// TIA Portal project "Pesteproject" (V15.1)

(* hardware
DEVICE "S7-1200 station_1"  S7-1200 Station
   slot 0: "Rack_0"  S7-1200 Rack  Rack  V1.0
   slot 1: "PLC_Lines_A_B"  CPU 1212C AC/DC/Rly  6ES7 212-1BE40-0XB0  V4.2
   slot 2: "DI 16x24VDC/DQ 16xRelay_1"  SM 1223 DI16/DQ16 x relay  6ES7 223-1PL32-0XB0  V2.0
   slot 3: "CB 1241 (RS485)"  CB 1241 (RS485)  6ES7 241-1CH30-1XB0  V1.0
   slot 3: "DQ 16xRelay_1"  SM 1222 DQ16 x relay  6ES7 222-1HH32-0XB0  V2.0
DEVICE "S7-1200 station_2"  S7-1200 Station
   slot 0: "Rack_0"  S7-1200 Rack  Rack  V1.0
   slot 1: "PLC_Lines_C"  CPU 1212C AC/DC/Rly  6ES7 212-1BE40-0XB0  V4.2
   slot 2: "DQ 16xRelay_1"  SM 1222 DQ16 x relay  6ES7 222-1HH32-0XB0  V2.0
   slot 3: "CB 1241 (RS485)"  CB 1241 (RS485)  6ES7 241-1CH30-1XB0  V1.0
DEVICE "S71500/ET200MP station_1"  S7-1500 station
   slot 0: "Rail_0"  Rack  6ES7 590-1***0-0AA0
   slot 1: "PLC_1"  CPU 1516-3 PN/DP  6ES7 516-3AN01-0AB0  V2.5
      slot 3: "CPU display_1"  6ES7591-1BA00-0AA0
   slot 2: "DI 16x24VDC BA_1"  DI 16x24VDC BA  6ES7 521-1BH10-0AA0  V1.1
   slot 3: "DI 16x24VDC BA_2"  DI 16x24VDC BA  6ES7 521-1BH10-0AA0  V1.1
*)

// ===== PLC "PLC_Lines_A_B"  CPU 1212C AC/DC/Rly =====

VAR_GLOBAL   // PLC tag table "Default tag table"
   "Phase_Control" AT %I8.0 : Bool;
   "Start_A" AT %I8.7 : Bool;
   "Spare_6" AT %I9.6 : Bool;
   "Spare_7" AT %I9.7 : Bool;
   "Emergency_A" AT %I8.4 : Bool;
   "Fault_A1" AT %I8.1 : Bool;
   "Low_Silo_A1" AT %I0.2 : Bool;
   "Low_Silo_A2" AT %I0.1 : Bool;
   "Low_Silo_B1" AT %I0.7 : Bool;
   "Low_Silo_B2" AT %I0.4 : Bool;
   "High_Silo_A1" AT %I0.3 : Bool;
   "High_Silo_A2" AT %I0.0 : Bool;
   "High_Silo_B1" AT %I0.6 : Bool;
   "High_Silo_B2" AT %I0.5 : Bool;
   "Fault_A2" AT %I9.1 : Bool;
   "Fault_B1" AT %I8.2 : Bool;
   "Fault_B2" AT %I9.2 : Bool;
   "Fault_A3" AT %I9.5 : Bool;
   "Fault_B3" AT %I9.4 : Bool;
   "Emergency_B" AT %I9.3 : Bool;
   "Rel Spare_4" AT %Q2.4 : Bool;
   "Rel Spare_5" AT %Q2.5 : Bool;
   "Rel Spare_6" AT %Q2.6 : Bool;
   "Rel Spare_7" AT %Q2.7 : Bool;
   "Rel Spare_8" AT %Q3.0 : Bool;
   "Rel Spare_9" AT %Q3.1 : Bool;
   "Rel Spare_10" AT %Q3.2 : Bool;
   "Rel Spare_11" AT %Q3.3 : Bool;
   "Rel Spare_12" AT %Q3.4 : Bool;
   "Rel Spare_13" AT %Q3.5 : Bool;
   "Rel Spare_14" AT %Q3.6 : Bool;
   "Rel Spare_15" AT %Q3.7 : Bool;
   "Light_A1" AT %Q2.3 : Bool;
   "Light_A2" AT %Q2.2 : Bool;
   "Light_B1" AT %Q2.1 : Bool;
   "Light_B2" AT %Q2.0 : Bool;
   "Conveyer_A1" AT %Q0.4 : Bool;
   "Conveyer_A2" AT %Q0.5 : Bool;
   "Conveyer_B1" AT %Q9.0 : Bool;
   "Conveyer_B2" AT %Q8.0 : Bool;
   "Pneumatic_A1" AT %Q9.1 : Bool;
   "Pneumatic_A2" AT %Q8.1 : Bool;
   "Pneumatic_B1" AT %Q8.2 : Bool;
   "Pneumatic_B2" AT %Q9.2 : Bool;
   "Conveyer_A3" AT %Q9.5 : Bool;
   "Conveyer_B3_Left" AT %Q9.6 : Bool;
   "Conveyer_B3_Right" AT %Q8.5 : Bool;
   "Tag_1" AT %M10.0 : Bool;
   "Tag_2" AT %M10.1 : Bool;
   "start" AT %M10.2 : Bool;
   "Tag_3" AT %M110.0 : Bool;
   "Tag_10" AT %M110.1 : Bool;
   "Tag_11" AT %M110.2 : Bool;
   "System_Byte" AT %MB1 : Byte;
   "FirstScan" AT %M1.0 : Bool;
   "DiagStatusUpdate" AT %M1.1 : Bool;
   "AlwaysTRUE" AT %M1.2 : Bool;
   "AlwaysFALSE" AT %M1.3 : Bool;
   "Clock_Byte" AT %MB0 : Byte;
   "Clock_10Hz" AT %M0.0 : Bool;
   "Clock_5Hz" AT %M0.1 : Bool;
   "Clock_2.5Hz" AT %M0.2 : Bool;
   "Clock_2Hz" AT %M0.3 : Bool;
   "Clock_1.25Hz" AT %M0.4 : Bool;
   "Clock_1Hz" AT %M0.5 : Bool;
   "Clock_0.625Hz" AT %M0.6 : Bool;
   "Clock_0.5Hz" AT %M0.7 : Bool;
   "Tag_12" AT %M120.1 : Bool;
   "Tag_13" AT %M120.0 : Bool;
   "Tag_14" AT %M120.2 : Bool;
   "Tag_15" AT %MW112 : Word;
   "Tag_16" AT %MW114 : Word;
   "Tag_17" AT %MW122 : Word;
   "Tag_18" AT %MW124 : Word;
   "Tag_4" AT %M1000.0 : Bool;
   "Tag_5" AT %M1000.1 : Bool;
   "Tag_6" AT %MW1002 : Word;
   "Tag_7" AT %M1000.4 : Bool;
   "Tag_8" AT %MW1004 : Word;
   "Tag_9" AT %M1010.0 : Bool;
   "Tag_19" AT %M1010.1 : Bool;
   "Tag_20" AT %M1010.2 : Bool;
   "Tag_21" AT %MW1012 : Word;
   "Tag_22" AT %M1010.4 : Bool;
   "Tag_23" AT %MW1014 : Word;
   "Tag_24" AT %M990.0 : Bool;
   "Tag_25" AT %M990.5 : Bool;
   "Line_A1_Start_Consent" AT %M150.0 : Bool;
   "Line_A1_Run_Consent" AT %M150.1 : Bool;
   "Line_A1_Conveyer_Timer" AT %M150.2 : Bool;
   "A1_Start_Conveyer" AT %M150.3 : Bool;
   "TriggerStartToggleMemory" AT %M150.4 : Bool;
   "Start_A1_Toggle" AT %M150.5 : Bool;
   "TriggerA1ToggleStop" AT %M150.6 : Bool;
   "Conveyer_A1_On" AT %M150.7 : Bool;
   "Conveyer_A1_Off" AT %M151.0 : Bool;
   "Line_A2_Start_Consent" AT %M160.0 : Bool;
   "Line_A2_Run_Consent" AT %M160.1 : Bool;
   "Line_A2_Conveyer_Timer" AT %M160.2 : Bool;
   "A2_Start_Conveyer" AT %M160.3 : Bool;
   "TriggerStopToggleMemoryA2" AT %M160.6 : Bool;
   "TriggerStartToggleMemoryA2" AT %M160.4 : Bool;
   "Start_A2_Toggle" AT %M160.5 : Bool;
   "Conveyer_A2_Off" AT %M161.0 : Bool;
   "Conveyer_A2_On" AT %M160.7 : Bool;
   "Line_B1_Start_Consent" AT %M170.0 : Bool;
   "Line_B1_Run_Consent" AT %M170.1 : Bool;
   "Line_B1_Conveyer_Timer" AT %M170.2 : Bool;
   "B1_Start_Conveyer" AT %M170.3 : Bool;
   "Start_B1_Toggle" AT %M170.5 : Bool;
   "TriggerStartToggleMemoryB1" AT %M170.4 : Bool;
   "TriggerB1ToggleStop" AT %M170.6 : Bool;
   "Conveyer_B1_Off" AT %M171.0 : Bool;
   "Conveyer_B1_On" AT %M170.7 : Bool;
   "Line_B2_Start_Consent" AT %M180.0 : Bool;
   "Line_B2_Run_Consent" AT %M180.1 : Bool;
   "B2_Start_Conveyer" AT %M180.3 : Bool;
   "Line_B2_Conveyer_Timer" AT %M180.2 : Bool;
   "Start_B2_Toggle" AT %M180.5 : Bool;
   "TriggerStartToggleMemoryB2" AT %M180.4 : Bool;
   "TriggerStopToggleMemoryB2" AT %M180.6 : Bool;
   "Conveyer_B2_Off" AT %M181.0 : Bool;
   "Conveyer_B2_On" AT %M180.7 : Bool;
   "Vibrator_A1_On" AT %M151.4 : Bool;
   "Vibrator_A2_On" AT %M161.4 : Bool;
   "Vibrator_B1_On" AT %M171.4 : Bool;
   "Vibrator_B2_On" AT %M181.4 : Bool;
   "A1_Sample_Triger" AT %M151.1 : Bool;
   "Conveyer_A1_OneShut" AT %M151.2 : Bool;
   "Tag_27" AT %M151.3 : Bool;
   "A2_Sample_Triger" AT %M161.1 : Bool;
   "Conveyer_A2_OneShut" AT %M161.2 : Bool;
   "B1_Sample_Triger" AT %M171.1 : Bool;
   "Conveyer_B1_OneShut" AT %M171.2 : Bool;
   "B2_Sample_Triger" AT %M181.1 : Bool;
   "Conveyer_B2_OneShut" AT %M181.2 : Bool;
   "B_Emergency_Flag" AT %M171.3 : Bool;
   "SiloAToggleStart" AT %M190.0 : Bool;
   "SiloBToggleStart" AT %M190.1 : Bool;
   "Conveyor_B3_Left" AT %M200.0 : Bool;
   "Conveyor_B3_Right" AT %M200.1 : Bool;
   "Silo_B_Not_Start_Timer" AT %M190.3 : Bool;
   "Silo_A_Not_Start_Timer" AT %M190.2 : Bool;
   "Conveyor_B3_Start" AT %M190.4 : Bool;
   "Conveyor_A1_Empty_line" AT %M151.5 : Bool;
   "Conveyor_A2_Empty_line" AT %M161.5 : Bool;
   "Conveyor_B1_Empty_line" AT %M171.5 : Bool;
   "Conveyor_B2_Empty_line" AT %M181.5 : Bool;
   "Tag_26" AT %MD156 : DInt;
   "Tag_28" AT %MD166 : DInt;
   "Tag_29" AT %MD176 : DInt;
   "Tag_30" AT %MD186 : DInt;
END_VAR

TYPE "tIMEDATATYPE"
VERSION : 0.1
   STRUCT
      HOUR : String;
      MINUTE : String;
      DAY : String;
      MONTH : String;
      YEAR : String;
   END_STRUCT;
END_TYPE

DATA_BLOCK "ScenarioData"   // DB1
{ S7_Optimized_Access := 'TRUE' }
VERSION : 0.1
   VAR
      DefaultScenario : Int := 1;
      Line_A1_Conveyer_on_Time_Scenario_A : DInt := 2;
      Line_A1_Conveyer_off_Time_Scenario_A : DInt := 3;
      Line_A1_Sampling_Time_Scenario_A : DInt := 4;
      Line_A1_Sampling_OpenTime_Scenario_A : DInt := 5;
      Line_A1_Feeder_Intensity_Scenario_A : Int := 6;
      Line_A1_Duration_Big_Silo_Off_Scenario_A : DInt := 7;
      Line_A1_Feeder_Delay_Before_Stop_Time_Scenario_A : DInt := 8;
      Line_A1_Feeder_Delay_After_Start_Time_Scenario_A : DInt := 9;
      Line_A1_Conveyer_on_Time_Scenario_B : DInt := 10;
      Line_A1_Conveyer_off_Time_Scenario_B : DInt := 11;
      Line_A1_Sampling_Time_Scenario_B : DInt := 12;
      Line_A1_Sampling_OpenTime_Scenario_B : DInt := 13;
      Line_A1_Feeder_Intensity_Scenario_B : Int := 14;
      Line_A1_Duration_Big_Silo_Off_Scenario_B : DInt := 15;
      Line_A1_Feeder_Delay_Before_Stop_Time_Scenario_B : DInt := 16;
      Line_A1_Feeder_Delay_After_Start_Time_Scenario_B : DInt := 17;
      Line_A1_Conveyer_on_Time_Scenario_C : DInt := 18;
      Line_A1_Conveyer_off_Time_Scenario_C : DInt := 19;
      Line_A1_Sampling_Time_Scenario_C : DInt := 20;
      Line_A1_Sampling_OpenTime_Scenario_C : DInt := 21;
      Line_A1_Feeder_Intensity_Scenario_C : Int := 22;
      Line_A1_Duration_Big_Silo_Off_Scenario_C : DInt := 23;
      Line_A1_Feeder_Delay_Before_Stop_Time_Scenario_C : DInt := 24;
      Line_A1_Feeder_Delay_After_Start_Time_Scenario_C : DInt := 25;
      Line_A1_Conveyer_on_Time_Scenario_E : DInt := 26;
      Line_A1_Conveyer_off_Time_Scenario_E : DInt := 27;
      Line_A1_Sampling_Time_Scenario_E : DInt := 28;
      Line_A1_Sampling_OpenTime_Scenario_E : DInt := 29;
      Line_A1_Feeder_Intensity_Scenario_E : Int := 30;
      Line_A1_Duration_Big_Silo_Off_Scenario_E : DInt := 31;
      Line_A1_Feeder_Delay_Before_Stop_Time_Scenario_E : DInt := 32;
      Line_A1_Feeder_Delay_After_Start_Time_Scenario_E : DInt := 33;
      Line_A1_Conveyer_on_Time_Scenario_D : DInt := 34;
      Line_A1_Conveyer_off_Time_Scenario_D : DInt := 35;
      Line_A1_Sampling_Time_Scenario_D : DInt := 36;
      Line_A1_Sampling_OpenTime_Scenario_D : DInt := 37;
      Line_A1_Feeder_Intensity_Scenario_D : Int := 38;
      Line_A1_Duration_Big_Silo_Off_Scenario_D : DInt := 39;
      Line_A1_Feeder_Delay_Before_Stop_Time_Scenario_D : DInt := 40;
      Line_A1_Feeder_Delay_After_Start_Time_Scenario_D : DInt := 41;
      Line_A2_Conveyer_on_Time_Scenario_A : DInt := 42;
      Line_A2_Conveyer_off_Time_Scenario_A : DInt := 43;
      Line_A2_Sampling_Time_Scenario_A : DInt := 44;
      Line_A2_Sampling_OpenTime_Scenario_A : DInt := 45;
      Line_A2_Feeder_Intensity_Scenario_A : Int := 46;
      Line_A2_Duration_Big_Silo_Off_Scenario_A : DInt := 47;
      Line_A2_Feeder_Delay_Before_Stop_Time_Scenario_A : DInt := 48;
      Line_A2_Feeder_Delay_After_Start_Time_Scenario_A : DInt := 49;
      Line_A2_Conveyer_on_Time_Scenario_B : DInt := 50;
      Line_A2_Conveyer_off_Time_Scenario_B : DInt := 51;
      Line_A2_Sampling_Time_Scenario_B : DInt := 52;
      Line_A2_Sampling_OpenTime_Scenario_B : DInt := 53;
      Line_A2_Feeder_Intensity_Scenario_B : Int := 54;
      Line_A2_Duration_Big_Silo_Off_Scenario_B : DInt := 55;
      Line_A2_Feeder_Delay_Before_Stop_Time_Scenario_B : DInt := 56;
      Line_A2_Feeder_Delay_After_Start_Time_Scenario_B : DInt := 57;
      Line_A2_Conveyer_on_Time_Scenario_C : DInt := 58;
      Line_A2_Conveyer_off_Time_Scenario_C : DInt := 59;
      Line_A2_Sampling_Time_Scenario_C : DInt := 60;
      Line_A2_Sampling_OpenTime_Scenario_C : DInt := 61;
      Line_A2_Feeder_Intensity_Scenario_C : Int := 62;
      Line_A2_Duration_Big_Silo_Off_Scenario_C : DInt := 63;
      Line_A2_Feeder_Delay_Before_Stop_Time_Scenario_C : DInt := 64;
      Line_A2_Feeder_Delay_After_Start_Time_Scenario_C : DInt := 65;
      Line_A2_Conveyer_on_Time_Scenario_E : DInt := 66;
      Line_A2_Conveyer_off_Time_Scenario_E : DInt := 67;
      Line_A2_Sampling_Time_Scenario_E : DInt := 68;
      Line_A2_Sampling_OpenTime_Scenario_E : DInt := 69;
      Line_A2_Feeder_Intensity_Scenario_E : Int := 70;
      Line_A2_Duration_Big_Silo_Off_Scenario_E : DInt := 71;
      Line_A2_Feeder_Delay_Before_Stop_Time_Scenario_E : DInt := 72;
      Line_A2_Feeder_Delay_After_Start_Time_Scenario_E : DInt := 73;
      Line_A2_Conveyer_on_Time_Scenario_D : DInt := 74;
      Line_A2_Conveyer_off_Time_Scenario_D : DInt := 75;
      Line_A2_Sampling_Time_Scenario_D : DInt := 76;
      Line_A2_Sampling_OpenTime_Scenario_D : DInt := 77;
      Line_A2_Feeder_Intensity_Scenario_D : Int := 78;
      Line_A2_Duration_Big_Silo_Off_Scenario_D : DInt := 79;
      Line_A2_Feeder_Delay_Before_Stop_Time_Scenario_D : DInt := 80;
      Line_A2_Feeder_Delay_After_Start_Time_Scenario_D : DInt := 81;
      Line_B1_Conveyer_on_Time_Scenario_A : DInt := 82;
      Line_B1_Conveyer_off_Time_Scenario_A : DInt := 83;
      Line_B1_Sampling_Time_Scenario_A : DInt := 84;
      Line_B1_Sampling_OpenTime_Scenario_A : DInt := 85;
      Line_B1_Feeder_Intensity_Scenario_A : Int := 86;
      Line_B1_Duration_Big_Silo_Off_Scenario_A : DInt := 87;
      Line_B1_Feeder_Delay_Before_Stop_Time_Scenario_A : DInt := 88;
      Line_B1_Feeder_Delay_After_Start_Time_Scenario_A : DInt := 89;
      Line_B1_Conveyer_on_Time_Scenario_B : DInt := 90;
      Line_B1_Conveyer_off_Time_Scenario_B : DInt := 91;
      Line_B1_Sampling_Time_Scenario_B : DInt := 92;
      Line_B1_Sampling_OpenTime_Scenario_B : DInt := 93;
      Line_B1_Feeder_Intensity_Scenario_B : Int := 94;
      Line_B1_Duration_Big_Silo_Off_Scenario_B : DInt := 95;
      Line_B1_Feeder_Delay_Before_Stop_Time_Scenario_B : DInt := 96;
      Line_B1_Feeder_Delay_After_Start_Time_Scenario_B : DInt := 97;
      Line_B1_Conveyer_on_Time_Scenario_C : DInt := 98;
      Line_B1_Conveyer_off_Time_Scenario_C : DInt := 99;
      Line_B1_Sampling_Time_Scenario_C : DInt := 100;
      Line_B1_Sampling_OpenTime_Scenario_C : DInt := 101;
      Line_B1_Feeder_Intensity_Scenario_C : Int := 102;
      Line_B1_Duration_Big_Silo_Off_Scenario_C : DInt := 103;
      Line_B1_Feeder_Delay_Before_Stop_Time_Scenario_C : DInt := 104;
      Line_B1_Feeder_Delay_After_Start_Time_Scenario_C : DInt := 105;
      Line_B1_Conveyer_on_Time_Scenario_E : DInt := 106;
      Line_B1_Conveyer_off_Time_Scenario_E : DInt := 107;
      Line_B1_Sampling_Time_Scenario_E : DInt := 108;
      Line_B1_Sampling_OpenTime_Scenario_E : DInt := 109;
      Line_B1_Feeder_Intensity_Scenario_E : Int := 110;
      Line_B1_Duration_Big_Silo_Off_Scenario_E : DInt := 111;
      Line_B1_Feeder_Delay_Before_Stop_Time_Scenario_E : DInt := 112;
      Line_B1_Feeder_Delay_After_Start_Time_Scenario_E : DInt := 113;
      Line_B1_Conveyer_on_Time_Scenario_D : DInt := 114;
      Line_B1_Conveyer_off_Time_Scenario_D : DInt := 115;
      Line_B1_Sampling_Time_Scenario_D : DInt := 116;
      Line_B1_Sampling_OpenTime_Scenario_D : DInt := 117;
      Line_B1_Feeder_Intensity_Scenario_D : Int := 118;
      Line_B1_Duration_Big_Silo_Off_Scenario_D : DInt := 119;
      Line_B1_Feeder_Delay_Before_Stop_Time_Scenario_D : DInt := 120;
      Line_B1_Feeder_Delay_After_Start_Time_Scenario_D : DInt := 121;
      Line_B2_Conveyer_on_Time_Scenario_A : DInt := 122;
      Line_B2_Conveyer_off_Time_Scenario_A : DInt := 123;
      Line_B2_Sampling_Time_Scenario_A : DInt := 124;
      Line_B2_Sampling_OpenTime_Scenario_A : DInt := 125;
      Line_B2_Feeder_Intensity_Scenario_A : Int := 126;
      Line_B2_Duration_Big_Silo_Off_Scenario_A : DInt := 127;
      Line_B2_Feeder_Delay_Before_Stop_Time_Scenario_A : DInt := 128;
      Line_B2_Feeder_Delay_After_Start_Time_Scenario_A : DInt := 129;
      Line_B2_Conveyer_on_Time_Scenario_B : DInt := 130;
      Line_B2_Conveyer_off_Time_Scenario_B : DInt := 131;
      Line_B2_Sampling_Time_Scenario_B : DInt := 132;
      Line_B2_Sampling_OpenTime_Scenario_B : DInt := 133;
      Line_B2_Feeder_Intensity_Scenario_B : Int := 134;
      Line_B2_Duration_Big_Silo_Off_Scenario_B : DInt := 135;
      Line_B2_Feeder_Delay_Before_Stop_Time_Scenario_B : DInt := 136;
      Line_B2_Feeder_Delay_After_Start_Time_Scenario_B : DInt := 137;
      Line_B2_Conveyer_on_Time_Scenario_C : DInt := 138;
      Line_B2_Conveyer_off_Time_Scenario_C : DInt := 139;
      Line_B2_Sampling_Time_Scenario_C : DInt := 140;
      Line_B2_Sampling_OpenTime_Scenario_C : DInt := 141;
      Line_B2_Feeder_Intensity_Scenario_C : Int := 142;
      Line_B2_Duration_Big_Silo_Off_Scenario_C : DInt := 143;
      Line_B2_Feeder_Delay_Before_Stop_Time_Scenario_C : DInt := 144;
      Line_B2_Feeder_Delay_After_Start_Time_Scenario_C : DInt := 145;
      Line_B2_Conveyer_on_Time_Scenario_E : DInt := 146;
      Line_B2_Conveyer_off_Time_Scenario_E : DInt := 147;
      Line_B2_Sampling_Time_Scenario_E : DInt := 148;
      Line_B2_Sampling_OpenTime_Scenario_E : DInt := 149;
      Line_B2_Feeder_Intensity_Scenario_E : Int := 150;
      Line_B2_Duration_Big_Silo_Off_Scenario_E : DInt := 151;
      Line_B2_Feeder_Delay_Before_Stop_Time_Scenario_E : DInt := 152;
      Line_B2_Feeder_Delay_After_Start_Time_Scenario_E : DInt := 153;
      Line_B2_Conveyer_on_Time_Scenario_D : DInt := 154;
      Line_B2_Conveyer_off_Time_Scenario_D : DInt := 155;
      Line_B2_Sampling_Time_Scenario_D : DInt := 156;
      Line_B2_Sampling_OpenTime_Scenario_D : DInt := 157;
      Line_B2_Feeder_Intensity_Scenario_D : Int := 158;
      Line_B2_Duration_Big_Silo_Off_Scenario_D : DInt := 159;
      Line_B2_Feeder_Delay_Before_Stop_Time_Scenario_D : DInt := 160;
      Line_B2_Feeder_Delay_After_Start_Time_Scenario_D : DInt := 161;
      Line_A1_Empty_Line_Time_Scenario_A : DInt := 162;
      Line_A2_Empty_Line_Time_Scenario_A : DInt := 163;
      Line_B1_Empty_Line_Time_Scenario_A : DInt := 164;
      Line_B2_Empty_Line_Time_Scenario_A : DInt := 165;
      Line_A1_Empty_Line_Time_Scenario_B : DInt := 166;
      Line_A2_Empty_Line_Time_Scenario_B : DInt := 167;
      Line_B1_Empty_Line_Time_Scenario_B : DInt := 168;
      Line_B2_Empty_Line_Time_Scenario_B : DInt := 169;
      Line_A1_Empty_Line_Time_Scenario_C : DInt := 170;
      Line_A2_Empty_Line_Time_Scenario_C : DInt := 171;
      Line_B1_Empty_Line_Time_Scenario_C : DInt := 172;
      Line_B2_Empty_Line_Time_Scenario_C : DInt := 173;
      Line_A1_Empty_Line_Time_Scenario_D : DInt := 174;
      Line_A2_Empty_Line_Time_Scenario_D : DInt := 175;
      Line_B1_Empty_Line_Time_Scenario_D : DInt := 176;
      Line_B2_Empty_Line_Time_Scenario_D : DInt := 177;
      Line_A1_Empty_Line_Time_Scenario_E : DInt := 178;
      Line_A2_Empty_Line_Time_Scenario_E : DInt := 179;
      Line_B1_Empty_Line_Time_Scenario_E : DInt := 180;
      Line_B2_Empty_Line_Time_Scenario_E : DInt := 181;
   END_VAR
BEGIN
END_DATA_BLOCK

DATA_BLOCK "Conveyer B1_DB"   // DB5
{ S7_Optimized_Access := 'TRUE' }
VERSION : 0.1
// stored: InstanceOfName Conveyer B1
"Conveyer B1"
BEGIN
END_DATA_BLOCK

DATA_BLOCK "ModbusDataSendToFeeders"   // DB7
{ S7_Optimized_Access := 'FALSE' }
VERSION : 0.1
   VAR
      dataforsend : Array[0..3] of Int;
   END_VAR
BEGIN
   dataforsend[0] := 0;
   dataforsend[1] := 0;
   dataforsend[2] := 0;
   dataforsend[3] := 0;
END_DATA_BLOCK

DATA_BLOCK "Conveyer A1_DB"   // DB12
{ S7_Optimized_Access := 'TRUE' }
VERSION : 0.1
// stored: InstanceOfName Conveyer A1
"Conveyer A1"
BEGIN
END_DATA_BLOCK

DATA_BLOCK "Conveyer A2_DB"   // DB13
{ S7_Optimized_Access := 'TRUE' }
VERSION : 0.1
// stored: InstanceOfName Conveyer A2
"Conveyer A2"
BEGIN
END_DATA_BLOCK

DATA_BLOCK "Conveyer B1_DB_1"   // DB17
{ S7_Optimized_Access := 'TRUE' }
VERSION : 0.1
// stored: InstanceOfName Conveyer B1
"Conveyer B1"
BEGIN
END_DATA_BLOCK

DATA_BLOCK "Conveyer B2_DB"   // DB18
{ S7_Optimized_Access := 'TRUE' }
VERSION : 0.1
// stored: InstanceOfName Conveyer B2
"Conveyer B2"
BEGIN
END_DATA_BLOCK

DATA_BLOCK "Vibrator A1_DB"   // DB19
{ S7_Optimized_Access := 'TRUE' }
VERSION : 0.1
// stored: InstanceOfName Vibrator A1
"Vibrator A1"
BEGIN
END_DATA_BLOCK

DATA_BLOCK "Vibrator A2_DB"   // DB20
{ S7_Optimized_Access := 'TRUE' }
VERSION : 0.1
// stored: InstanceOfName Vibrator A2
"Vibrator A2"
BEGIN
END_DATA_BLOCK

DATA_BLOCK "Vibrator B1_DB"   // DB21
{ S7_Optimized_Access := 'TRUE' }
VERSION : 0.1
// stored: InstanceOfName Vibrator B1
"Vibrator B1"
BEGIN
END_DATA_BLOCK

DATA_BLOCK "Vibrator B2_DB"   // DB22
{ S7_Optimized_Access := 'TRUE' }
VERSION : 0.1
// stored: InstanceOfName Vibrator B2
"Vibrator B2"
BEGIN
END_DATA_BLOCK

DATA_BLOCK "Web_Send"   // DB23
{ S7_Optimized_Access := 'TRUE' }
VERSION : 0.1
   VAR
      "time" : DTL;
      ModbusDone : Bool;
      ModbusStatus : Word;
      A1_Scenario_Type : Int := 2;
      A2_Scenario_Type : Int := 1;
      B1_Scenario_Type : Int := 1;
      B2_Scenario_Type : Int := 1;
      A_Emergency : Bool;
      B_Emergency : Bool;
      A1_Fault : Bool;
      A2_Fault : Bool;
      B1_Fault : Bool;
      B2_Fault : Bool;
      A3_Fault : Bool;
      B3_Fault : Bool;
      A1_Silo_Low : Bool;
      A2_Silo_Low : Bool;
      B1_Silo_Low : Bool;
      B2_Silo_Low : Bool;
      A1_Conveyer : Bool;
      A2_Conveyer : Bool;
      B1_Conveyer : Bool;
      B2_Conveyer : Bool;
      A3_Conveyor : Bool;
      B3_Left_Conveyer : Bool;
      A1_Silo_High : Bool;
      A2_Silo_High : Bool;
      B1_Silo_High : Bool;
      B2_Silo_High : Bool;
      A1_Sample : Bool;
      A2_Sample : Bool;
      B1_Sample : Bool;
      B2_Sample : Bool;
      A1_Running_Duration : Time;
      A1_Pause_Duration : Time;
      A1_Feeder_Vibration_Intensity : Int;
      A1_Ruuning_Online : Time;
      A1_Pause_Online : Time;
      A1_Sample_Interval : Time;
      A1_Sample_Duration : Time;
      A1_Sample_Online : Time;
      A1_Enable : Bool;
      A1_Start : Bool;
      A1_Big_Silo : Bool;
      B1_Running_Duration : Time;
      B1_Pause_Duration : Time;
      B1_Feeder_Vibration_Intensity : Int;
      B1_Ruuning_Online : Time;
      B1_Pause_Online : Time;
      B1_Sample_Interval : Time;
      B1_Sample_Duration : Time;
      B1_Sample_Online : Time;
      B1_Enable : Bool;
      B1_Start : Bool;
      B1_Big_Silo : Bool;
      A2_Running_Duration : Time;
      A2_Pause_Duration : Time;
      A2_Feeder_Vibration_Intensity : Int;
      A2_Ruuning_Online : Time;
      A2_Pause_Online : Time;
      A2_Sample_Interval : Time;
      A2_Sample_Duration : Time;
      A2_Sample_Online : Time;
      A2_Enable : Bool;
      A2_Start : Bool;
      A2_Big_Silo : Bool;
      B2_Running_Duration : Time;
      B2_Pause_Duration : Time;
      B2_Feeder_Vibration_Intensity : Int;
      B2_Ruuning_Online : Time;
      B2_Pause_Online : Time;
      B2_Sample_Interval : Time;
      B2_Sample_Duration : Time;
      B2_Sample_Online : Time;
      B2_Enable : Bool;
      B2_Start : Bool;
      B2_Big_Silo : Bool;
      A1_Manual : Bool;
      A2_Manual : Bool;
      B1_Manual : Bool;
      B2_Manual : Bool;
      A1_Feeder : Bool;
      A2_Feeder : Bool;
      B1_Feeder : Bool;
      B2_Feeder : Bool;
      A1_Duration_Big_Silo_Stop_Time : Time;
      A2_Duration_Big_Silo_Stop_Time : Time;
      B1_Duration_Big_Silo_Stop_Time : Time;
      B2_Duration_Big_Silo_Stop_Time : Time;
      A1_Empty_Line_Time : Time;
      A2_Empty_Line_Time : Time;
      B1_Empty_Line_Time : Time;
      B2_Empty_Line_Time : Time;
      A1_Feeder_Delay_After_Start_Time : Time;
      A2_Feeder_Delay_After_Start_Time : Time;
      B1_Feeder_Delay_After_Start_Time : Time;
      B2_Feeder_Delay_After_Start_Time : Time;
      A1_Feeder_Delay_Before_Stop_Time : Time;
      A2_Feeder_Delay_Before_Stop_Time : Time;
      B1_Feeder_Delay_Before_Stop_Time : Time;
      B2_Feeder_Delay_Before_Stop_Time : Time;
      A1_Feeder_Delay_Time : Time;
      A1_Feeder_Delay_Time_1 : Time;
      A1_Feeder_Delay_Time_2 : Time;
      A1_Feeder_Delay_Time_3 : Time;
      B3_Conveyor : Bool;
   END_VAR
BEGIN
END_DATA_BLOCK

DATA_BLOCK "ConveyerA3_B3_DB"   // DB32
{ S7_Optimized_Access := 'TRUE' }
VERSION : 0.1
// stored: InstanceOfName ConveyerA3_B3
"ConveyerA3_B3"
BEGIN
END_DATA_BLOCK

DATA_BLOCK "Sample_A_DB"   // DB33
{ S7_Optimized_Access := 'TRUE' }
VERSION : 0.1
// stored: InstanceOfName Sample
"Sample"
BEGIN
END_DATA_BLOCK

DATA_BLOCK "Silo_Big_A-B_DB"   // DB34
{ S7_Optimized_Access := 'TRUE' }
VERSION : 0.1
// stored: InstanceOfName Silo_Big_A-B
"Silo_Big_A-B"
BEGIN
END_DATA_BLOCK

DATA_BLOCK "Web_Recieve"   // DB45
{ S7_Optimized_Access := 'FALSE' }
VERSION : 0.1
   VAR
      Line_A1_Save_Data : Bool;
      Line_A1_Save_Data_Advance : Bool;
      Line_A1_Start : Bool;
      Line_A1_Enable : Bool := 0;
      Line_A1_Conveyer_on_Time : Time := T#26MS;
      Line_A1_Conveyer_off_Time : Time := T#27MS;
      Line_A1_Sampling_Time : Time := T#28MS;
      Line_A1_Sampling_OpenTime : Time := T#29MS;
      Line_A1_Feeder_Intensity : Int := 30;
      Line_A1_Feeder_DelayTime : Time;
      Line_A1_Enable_Manual : Bool;
      Line_A1_Conveyor_Start_Manual : Bool;
      Line_A1_Big_Silo_Start_Manual : Bool;
      Line_A1_Below_Conveyor_Start_Manual : Bool;
      Line_A1_Feeder_Start_Manual : Bool;
      Line_A1_Sample_Start_Manual : Bool;
      Line_A1_Feeder_Delay_Before_Stop_Time : Time;
      Line_A1_Empty_Line_Time : Time;
      Line_A1_Big_Silo_Delay_Start : Time;
      Line_A1_Empty_Line : Bool;
      Line_A1_Feeder_Delay_After_Start_Time : Time;
      Line_A2_Save_Data : Bool;
      Line_A2_Save_Data_Advance : Bool;
      Line_A2_Start : Bool;
      Line_A2_Enable : Bool;
      Line_A2_Conveyer_on_Time : Time := T#8S_400MS;
      Line_A2_Conveyer_off_Time : Time := T#30s;
      Line_A2_Sampling_Time : Time := T#2M;
      Line_A2_Sampling_OpenTime : Time := T#9S_500MS;
      Line_A2_Feeder_Intensity : Int;
      Line_A2_Feeder_DelayTime : Time;
      Line_A2_Enable_Manual : Bool;
      Line_A2_Conveyor_Start_Manual : Bool;
      Line_A2_Big_Silo_Start_Manual : Bool;
      Line_A2_Below_Conveyor_Start_Manual : Bool;
      Line_A2_Feeder_Start_Manual : Bool;
      Line_A2_Sample_Start_Manual : Bool;
      Line_A2_Feeder_Delay_Before_Stop_Time : Time;
      Line_A2_Empty_Line_Time : Time;
      Line_A2_Big_Silo_Delay_Start : Time;
      Line_A2_Empty_Line : Bool;
      Line_A2_Feeder_Delay_After_Start_Time : Time;
      Line_B1_Save_Data : Bool;
      Line_B1_Save_Data_Advance : Bool;
      Line_B1_Start : Bool;
      Line_B1_Enable : Bool := 0;
      Line_B1_Conveyer_on_Time : Time := T#8S_400MS;
      Line_B1_Conveyer_off_Time : Time := T#30s;
      Line_B1_Sampling_Time : Time := T#2M;
      Line_B1_Sampling_OpenTime : Time := T#9S_500MS;
      Line_B1_Feeder_Intensity : Int;
      Line_B1_Feeder_DelayTime : Time;
      Line_B1_Enable_Manual : Bool;
      Line_B1_Conveyor_Start_Manual : Bool;
      Line_B1_Big_Silo_Start_Manual : Bool;
      Line_B1_Below_Conveyor_Start_Manual : Bool;
      Line_B1_Feeder_Start_Manual : Bool;
      Line_B1_Sample_Start_Manual : Bool;
      Line_B1_Feeder_Delay_Before_Stop_Time : Time;
      Line_B1_Empty_Line_Time : Time;
      Line_B1_Big_Silo_Delay_Start : Time;
      Line_B1_Empty_Line : Bool;
      Line_B1_Feeder_Delay_After_Start_Time : Time;
      Line_B2_Save_Data : Bool;
      Line_B2_Save_Data_Advance : Bool;
      Line_B2_Start : Bool;
      Line_B2_Enable : Bool := 0;
      Line_B2_Conveyer_on_Time : Time := T#8S_400MS;
      Line_B2_Conveyer_off_Time : Time := T#30s;
      Line_B2_Sampling_Time : Time := T#2M;
      Line_B2_Sampling_OpenTime : Time := T#9S_500MS;
      Line_B2_Feeder_Intensity : Int;
      Line_B2_Feeder_DelayTime : Time;
      Line_B2_Enable_Manual : Bool;
      Line_B2_Conveyor_Start_Manual : Bool;
      Line_B2_Big_Silo_Start_Manual : Bool;
      Line_B2_Below_Conveyor_Start_Manual : Bool;
      Line_B2_Feeder_Start_Manual : Bool;
      Line_B2_Sample_Start_Manual : Bool;
      Line_B2_Feeder_Delay_Before_Stop_Time : Time;
      Line_B2_Empty_Line_Time : Time;
      Line_B2_Big_Silo_Delay_Start : Time;
      Line_B2_Empty_Line : Bool;
      Line_B2_Feeder_Delay_After_Start_Time : Time;
      Conveyer_B3_Left : Bool;
   END_VAR
BEGIN
END_DATA_BLOCK

DATA_BLOCK "Empty Line A1 A2_DB"   // DB47
{ S7_Optimized_Access := 'TRUE' }
VERSION : 0.1
// stored: InstanceOfName Empty Line A1 A2
"Empty Line A1 A2"
BEGIN
END_DATA_BLOCK

DATA_BLOCK "Empty Line B1 B2_DB"   // DB48
{ S7_Optimized_Access := 'TRUE' }
VERSION : 0.1
// stored: InstanceOfName Empty Line B1 B2
"Empty Line B1 B2"
BEGIN
END_DATA_BLOCK

DATA_BLOCK "WebDataPrepaare_DB"   // DB49
{ S7_Optimized_Access := 'TRUE' }
VERSION : 0.1
// stored: InstanceOfName WebDataPrepaare
"WebDataPrepaare"
BEGIN
END_DATA_BLOCK

DATA_BLOCK "SaveDataToDataBlock A1_DB"   // DB51
{ S7_Optimized_Access := 'TRUE' }
VERSION : 0.1
// stored: InstanceOfName SaveDataToDataBlock A1
"SaveDataToDataBlock A1"
BEGIN
END_DATA_BLOCK

DATA_BLOCK "SaveDataToDataBlock A2_DB"   // DB52
{ S7_Optimized_Access := 'TRUE' }
VERSION : 0.1
// stored: InstanceOfName SaveDataToDataBlock A2
"SaveDataToDataBlock A2"
BEGIN
END_DATA_BLOCK

DATA_BLOCK "SaveDataToDataBlock B1_DB"   // DB53
{ S7_Optimized_Access := 'TRUE' }
VERSION : 0.1
// stored: InstanceOfName SaveDataToDataBlock B1
"SaveDataToDataBlock B1"
BEGIN
END_DATA_BLOCK

DATA_BLOCK "SaveDataToDataBlock B2_DB"   // DB54
{ S7_Optimized_Access := 'TRUE' }
VERSION : 0.1
// stored: InstanceOfName SaveDataToDataBlock B2
"SaveDataToDataBlock B2"
BEGIN
END_DATA_BLOCK

// folder: System blocks/Program resources

DATA_BLOCK "Timer_On_B1_Conveyer"   // DB2
{ S7_Optimized_Access := 'TRUE' }
AUTHOR : Simatic
FAMILY : IEC
NAME : IEC_TMR
VERSION : 1.0
// stored: InstanceOfName IEC_TIMER
"IEC_TIMER"
BEGIN
END_DATA_BLOCK

DATA_BLOCK "Timer_On_A1_Conveyer"   // DB6
{ S7_Optimized_Access := 'TRUE' }
AUTHOR : Simatic
FAMILY : IEC
NAME : IEC_TMR
VERSION : 1.0
// stored: InstanceOfName IEC_TIMER
"IEC_TIMER"
BEGIN
END_DATA_BLOCK

DATA_BLOCK "Timer_Off_A1_Conveyer"   // DB8
{ S7_Optimized_Access := 'TRUE' }
AUTHOR : Simatic
FAMILY : IEC
NAME : IEC_TMR
VERSION : 1.0
// stored: InstanceOfName IEC_TIMER
"IEC_TIMER"
BEGIN
END_DATA_BLOCK

DATA_BLOCK "Timer_On_A2_Conveyer"   // DB10
{ S7_Optimized_Access := 'TRUE' }
AUTHOR : Simatic
FAMILY : IEC
NAME : IEC_TMR
VERSION : 1.0
// stored: InstanceOfName IEC_TIMER
"IEC_TIMER"
BEGIN
END_DATA_BLOCK

DATA_BLOCK "Timer_Off_A2_Conveyer"   // DB11
{ S7_Optimized_Access := 'TRUE' }
AUTHOR : Simatic
FAMILY : IEC
NAME : IEC_TMR
VERSION : 1.0
// stored: InstanceOfName IEC_TIMER
"IEC_TIMER"
BEGIN
END_DATA_BLOCK

DATA_BLOCK "Timer_Off_B1_Conveyer"   // DB14
{ S7_Optimized_Access := 'TRUE' }
AUTHOR : Simatic
FAMILY : IEC
NAME : IEC_TMR
VERSION : 1.0
// stored: InstanceOfName IEC_TIMER
"IEC_TIMER"
BEGIN
END_DATA_BLOCK

DATA_BLOCK "Timer_On_B2_Conveyer"   // DB15
{ S7_Optimized_Access := 'TRUE' }
AUTHOR : Simatic
FAMILY : IEC
NAME : IEC_TMR
VERSION : 1.0
// stored: InstanceOfName IEC_TIMER
"IEC_TIMER"
BEGIN
END_DATA_BLOCK

DATA_BLOCK "Timer_Off_B2_Conveyer"   // DB16
{ S7_Optimized_Access := 'TRUE' }
AUTHOR : Simatic
FAMILY : IEC
NAME : IEC_TMR
VERSION : 1.0
// stored: InstanceOfName IEC_TIMER
"IEC_TIMER"
BEGIN
END_DATA_BLOCK

DATA_BLOCK "Timer_Before_On_Sample_A1"   // DB24
{ S7_Optimized_Access := 'TRUE' }
AUTHOR : Simatic
FAMILY : IEC
NAME : IEC_TMR
VERSION : 1.0
// stored: InstanceOfName IEC_TIMER
"IEC_TIMER"
BEGIN
END_DATA_BLOCK

DATA_BLOCK "Timer_Sample_Open_Time_A1"   // DB25
{ S7_Optimized_Access := 'TRUE' }
AUTHOR : Simatic
FAMILY : IEC
NAME : IEC_TMR
VERSION : 1.0
// stored: InstanceOfName IEC_TIMER
"IEC_TIMER"
BEGIN
END_DATA_BLOCK

DATA_BLOCK "Timer_Before_On_Sample_A2"   // DB26
{ S7_Optimized_Access := 'TRUE' }
AUTHOR : Simatic
FAMILY : IEC
NAME : IEC_TMR
VERSION : 1.0
// stored: InstanceOfName IEC_TIMER
"IEC_TIMER"
BEGIN
END_DATA_BLOCK

DATA_BLOCK "Timer_Before_On_Sample_B1"   // DB27
{ S7_Optimized_Access := 'TRUE' }
AUTHOR : Simatic
FAMILY : IEC
NAME : IEC_TMR
VERSION : 1.0
// stored: InstanceOfName IEC_TIMER
"IEC_TIMER"
BEGIN
END_DATA_BLOCK

DATA_BLOCK "Timer_Sample_Open_Time_B1"   // DB28
{ S7_Optimized_Access := 'TRUE' }
AUTHOR : Simatic
FAMILY : IEC
NAME : IEC_TMR
VERSION : 1.0
// stored: InstanceOfName IEC_TIMER
"IEC_TIMER"
BEGIN
END_DATA_BLOCK

DATA_BLOCK "Timer_Before_On_Sample_B2"   // DB29
{ S7_Optimized_Access := 'TRUE' }
AUTHOR : Simatic
FAMILY : IEC
NAME : IEC_TMR
VERSION : 1.0
// stored: InstanceOfName IEC_TIMER
"IEC_TIMER"
BEGIN
END_DATA_BLOCK

DATA_BLOCK "Timer_Sample_Open_Time_B2"   // DB30
{ S7_Optimized_Access := 'TRUE' }
AUTHOR : Simatic
FAMILY : IEC
NAME : IEC_TMR
VERSION : 1.0
// stored: InstanceOfName IEC_TIMER
"IEC_TIMER"
BEGIN
END_DATA_BLOCK

DATA_BLOCK "Timer_Sample_Open_Time_A2"   // DB31
{ S7_Optimized_Access := 'TRUE' }
AUTHOR : Simatic
FAMILY : IEC
NAME : IEC_TMR
VERSION : 1.0
// stored: InstanceOfName IEC_TIMER
"IEC_TIMER"
BEGIN
END_DATA_BLOCK

DATA_BLOCK "Timer_Silo_Big_B_Off_Time"   // DB36
{ S7_Optimized_Access := 'TRUE' }
AUTHOR : Simatic
FAMILY : IEC
NAME : IEC_TMR
VERSION : 1.0
// stored: InstanceOfName IEC_TIMER
"IEC_TIMER"
BEGIN
END_DATA_BLOCK

DATA_BLOCK "Timer_Silo_Big_A_Off_Time"   // DB37
{ S7_Optimized_Access := 'TRUE' }
AUTHOR : Simatic
FAMILY : IEC
NAME : IEC_TMR
VERSION : 1.0
// stored: InstanceOfName IEC_TIMER
"IEC_TIMER"
BEGIN
END_DATA_BLOCK

DATA_BLOCK "A1_Feeder_On_Delay_Timer"   // DB38
{ S7_Optimized_Access := 'TRUE' }
AUTHOR : Simatic
FAMILY : IEC
NAME : IEC_TMR
VERSION : 1.0
// stored: InstanceOfName IEC_TIMER
"IEC_TIMER"
BEGIN
END_DATA_BLOCK

DATA_BLOCK "A2_Feeder_On_Delay_Timer"   // DB39
{ S7_Optimized_Access := 'TRUE' }
AUTHOR : Simatic
FAMILY : IEC
NAME : IEC_TMR
VERSION : 1.0
// stored: InstanceOfName IEC_TIMER
"IEC_TIMER"
BEGIN
END_DATA_BLOCK

DATA_BLOCK "B1_Feeder_On_Delay_Timer"   // DB40
{ S7_Optimized_Access := 'TRUE' }
AUTHOR : Simatic
FAMILY : IEC
NAME : IEC_TMR
VERSION : 1.0
// stored: InstanceOfName IEC_TIMER
"IEC_TIMER"
BEGIN
END_DATA_BLOCK

DATA_BLOCK "B2_Feeder_On_Delay_Timer"   // DB41
{ S7_Optimized_Access := 'TRUE' }
AUTHOR : Simatic
FAMILY : IEC
NAME : IEC_TMR
VERSION : 1.0
// stored: InstanceOfName IEC_TIMER
"IEC_TIMER"
BEGIN
END_DATA_BLOCK

DATA_BLOCK "Timer_A1_Empty_Line_DB"   // DB42
{ S7_Optimized_Access := 'TRUE' }
AUTHOR : Simatic
FAMILY : IEC
NAME : IEC_TMR
VERSION : 1.0
// stored: InstanceOfName IEC_TIMER
"IEC_TIMER"
BEGIN
END_DATA_BLOCK

DATA_BLOCK "Timer_A2_Empty_Line_DB"   // DB43
{ S7_Optimized_Access := 'TRUE' }
AUTHOR : Simatic
FAMILY : IEC
NAME : IEC_TMR
VERSION : 1.0
// stored: InstanceOfName IEC_TIMER
"IEC_TIMER"
BEGIN
END_DATA_BLOCK

DATA_BLOCK "Timer_B1_Empty_Line_DB"   // DB44
{ S7_Optimized_Access := 'TRUE' }
AUTHOR : Simatic
FAMILY : IEC
NAME : IEC_TMR
VERSION : 1.0
// stored: InstanceOfName IEC_TIMER
"IEC_TIMER"
BEGIN
END_DATA_BLOCK

DATA_BLOCK "Timer_B2_Empty_Line_DB"   // DB46
{ S7_Optimized_Access := 'TRUE' }
AUTHOR : Simatic
FAMILY : IEC
NAME : IEC_TMR
VERSION : 1.0
// stored: InstanceOfName IEC_TIMER
"IEC_TIMER"
BEGIN
END_DATA_BLOCK

DATA_BLOCK "Timer_A1_Reset_Save_Data"   // DB50
{ S7_Optimized_Access := 'TRUE' }
AUTHOR : Simatic
FAMILY : IEC
NAME : IEC_TMR
VERSION : 1.0
// stored: InstanceOfName IEC_TIMER
"IEC_TIMER"
BEGIN
END_DATA_BLOCK

// folder: (top level)

FUNCTION_BLOCK "Conveyer A1"   // FB1, LAD
{ S7_Optimized_Access := 'TRUE' }
VERSION : 0.1
   VAR_TEMP   // added for the SCL form of the ladder/FBD networks
      _w1 : Bool;
      _w2 : Bool;
   END_VAR
BEGIN

REGION Network 1: Start Consent line A1
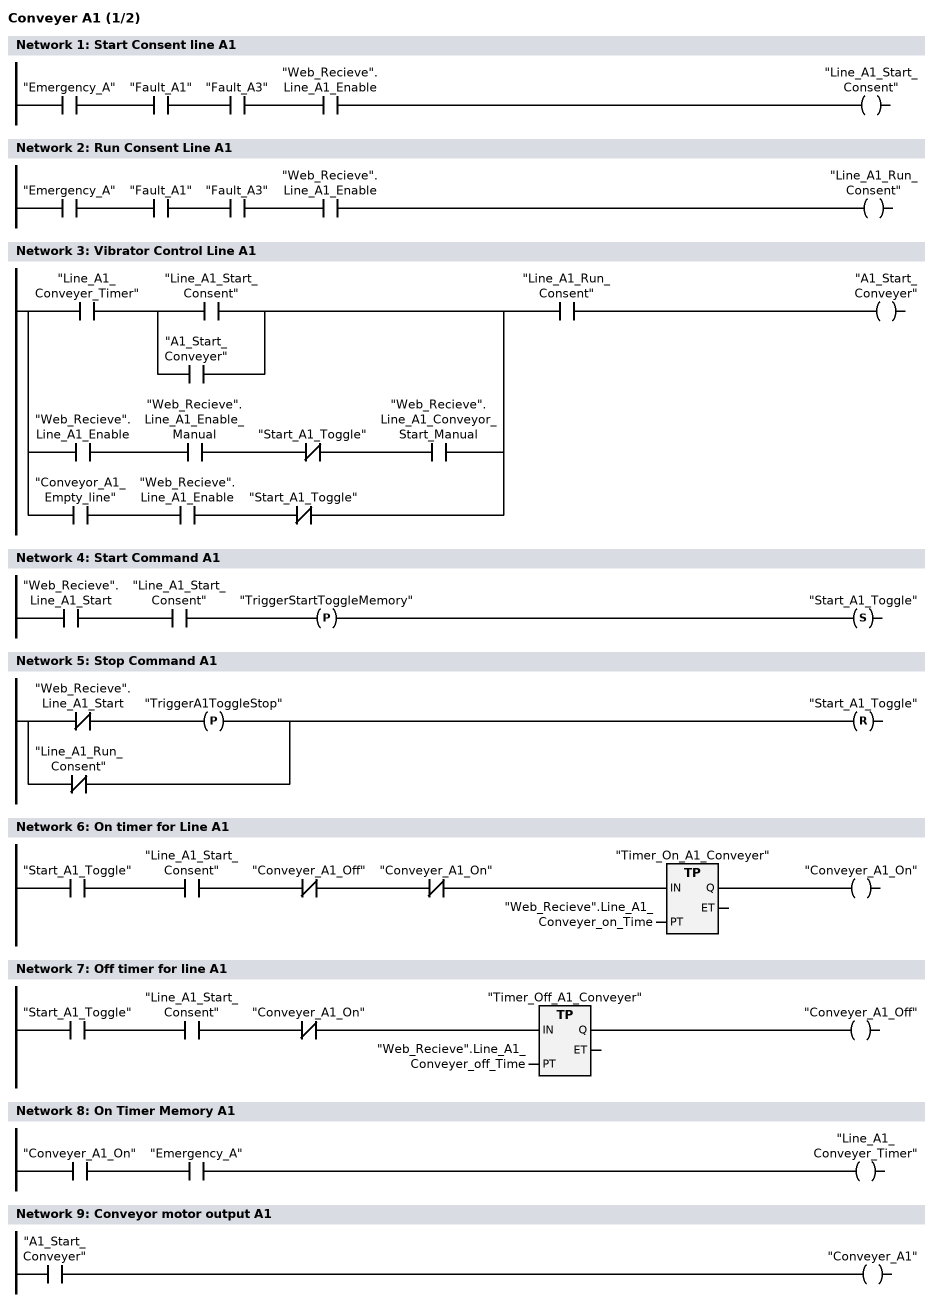
   RUNG wire#powerrail
      Contact( "Emergency_A" )
      Contact( "Fault_A1" )
      Contact( "Fault_A3" )
      Contact( "Web_Recieve".Line_A1_Enable )
      Coil( "Line_A1_Start_Consent" )
   END_RUNG
   // the same network as SCL:
   "Line_A1_Start_Consent" := "Emergency_A" AND "Fault_A1" AND "Fault_A3" AND "Web_Recieve".Line_A1_Enable;
END_REGION

REGION Network 2: Run Consent Line A1
   RUNG wire#powerrail
      Contact( "Emergency_A" )
      Contact( "Fault_A1" )
      Contact( "Fault_A3" )
      Contact( "Web_Recieve".Line_A1_Enable )
      Coil( "Line_A1_Run_Consent" )
   END_RUNG
   // the same network as SCL:
   "Line_A1_Run_Consent" := "Emergency_A" AND "Fault_A1" AND "Fault_A3" AND "Web_Recieve".Line_A1_Enable;
END_REGION

REGION Network 3: Vibrator Control Line A1
   RUNG wire#powerrail
      Contact( "Line_A1_Conveyer_Timer" )
      wire#w1
      Contact( "Line_A1_Start_Consent" )
      wire#w2
      Contact( "Line_A1_Run_Consent" )
      Coil( "A1_Start_Conveyer" )
   END_RUNG
   RUNG wire#w1
      Contact( "A1_Start_Conveyer" )
   END_RUNG wire#w2
   RUNG wire#powerrail
      Contact( "Web_Recieve".Line_A1_Enable )
      Contact( "Web_Recieve".Line_A1_Enable_Manual )
      I_Contact( "Start_A1_Toggle" )
      Contact( "Web_Recieve".Line_A1_Conveyor_Start_Manual )
   END_RUNG wire#w2
   RUNG wire#powerrail
      Contact( "Conveyor_A1_Empty_line" )
      Contact( "Web_Recieve".Line_A1_Enable )
      I_Contact( "Start_A1_Toggle" )
   END_RUNG wire#w2
   // the same network as SCL:
   "A1_Start_Conveyer" := (("Line_A1_Conveyer_Timer" AND ("Line_A1_Start_Consent" OR "A1_Start_Conveyer")) OR ("Web_Recieve".Line_A1_Enable AND "Web_Recieve".Line_A1_Enable_Manual AND NOT "Start_A1_Toggle" AND "Web_Recieve".Line_A1_Conveyor_Start_Manual) OR ("Conveyor_A1_Empty_line" AND "Web_Recieve".Line_A1_Enable AND NOT "Start_A1_Toggle")) AND "Line_A1_Run_Consent";
END_REGION

REGION Network 4: Start Command A1
   RUNG wire#powerrail
      Contact( "Web_Recieve".Line_A1_Start )
      Contact( "Line_A1_Start_Consent" )
      P_Trig( "TriggerStartToggleMemory" )
      S_Coil( "Start_A1_Toggle" )
   END_RUNG
   // the same network as SCL:
   #_w1 := "Web_Recieve".Line_A1_Start AND "Line_A1_Start_Consent";
   #_w2 := #_w1 AND NOT "TriggerStartToggleMemory";   // rising edge
   "TriggerStartToggleMemory" := #_w1;
   IF #_w2 THEN "Start_A1_Toggle" := TRUE; END_IF;
END_REGION

REGION Network 5: Stop Command A1
   RUNG wire#powerrail
      I_Contact( "Web_Recieve".Line_A1_Start )
      P_Trig( "TriggerA1ToggleStop" )
      wire#w1
      R_Coil( "Start_A1_Toggle" )
   END_RUNG
   RUNG wire#powerrail
      I_Contact( "Line_A1_Run_Consent" )
   END_RUNG wire#w1
   // the same network as SCL:
   #_w1 := NOT "Web_Recieve".Line_A1_Start AND NOT "TriggerA1ToggleStop";   // rising edge
   "TriggerA1ToggleStop" := NOT "Web_Recieve".Line_A1_Start;
   IF #_w1 OR NOT "Line_A1_Run_Consent" THEN "Start_A1_Toggle" := FALSE; END_IF;
END_REGION

REGION Network 6: On timer for Line A1
   "Timer_On_A1_Conveyer".TP(IN := "Start_A1_Toggle" AND "Line_A1_Start_Consent" AND NOT "Conveyer_A1_Off" AND NOT "Conveyer_A1_On",
                           PT := "Web_Recieve".Line_A1_Conveyer_on_Time);
   "Conveyer_A1_On" := "Timer_On_A1_Conveyer".Q;
END_REGION

REGION Network 7: Off timer for line A1
   "Timer_Off_A1_Conveyer".TP(IN := "Start_A1_Toggle" AND "Line_A1_Start_Consent" AND NOT "Conveyer_A1_On",
                           PT := "Web_Recieve".Line_A1_Conveyer_off_Time);
   "Conveyer_A1_Off" := "Timer_Off_A1_Conveyer".Q;
END_REGION

REGION Network 8: On Timer Memory A1
   RUNG wire#powerrail
      Contact( "Conveyer_A1_On" )
      Contact( "Emergency_A" )
      Coil( "Line_A1_Conveyer_Timer" )
   END_RUNG
   // the same network as SCL:
   "Line_A1_Conveyer_Timer" := "Conveyer_A1_On" AND "Emergency_A";
END_REGION

REGION Network 9: Conveyor motor output A1
   RUNG wire#powerrail
      Contact( "A1_Start_Conveyer" )
      Coil( "Conveyer_A1" )
   END_RUNG
   // the same network as SCL:
   "Conveyer_A1" := "A1_Start_Conveyer";
END_REGION

REGION Network 10: emergency or stop or disable reser Timers A1
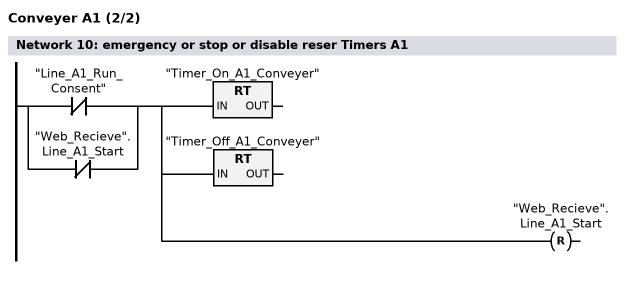
   RUNG wire#powerrail
      I_Contact( "Line_A1_Run_Consent" )
      wire#w1
      RT_Coil( "Timer_On_A1_Conveyer" )
   END_RUNG
   RUNG wire#powerrail
      I_Contact( "Web_Recieve".Line_A1_Start )
   END_RUNG wire#w1
   RUNG wire#w1
      RT_Coil( "Timer_Off_A1_Conveyer" )
   END_RUNG
   RUNG wire#w1
      R_Coil( "Web_Recieve".Line_A1_Start )
   END_RUNG
   // the same network as SCL:
   #_w1 := NOT "Line_A1_Run_Consent" OR NOT "Web_Recieve".Line_A1_Start;
   IF #_w1 THEN
       RESET_TIMER("Timer_On_A1_Conveyer");
       RESET_TIMER("Timer_Off_A1_Conveyer");
       "Web_Recieve".Line_A1_Start := FALSE;
   END_IF;
END_REGION
END_FUNCTION_BLOCK

FUNCTION_BLOCK "Conveyer A2"   // FB2, LAD
{ S7_Optimized_Access := 'TRUE' }
VERSION : 0.1
   VAR_TEMP   // added for the SCL form of the ladder/FBD networks
      _w1 : Bool;
      _w2 : Bool;
   END_VAR
BEGIN

REGION Network 1: Start Consent line A1